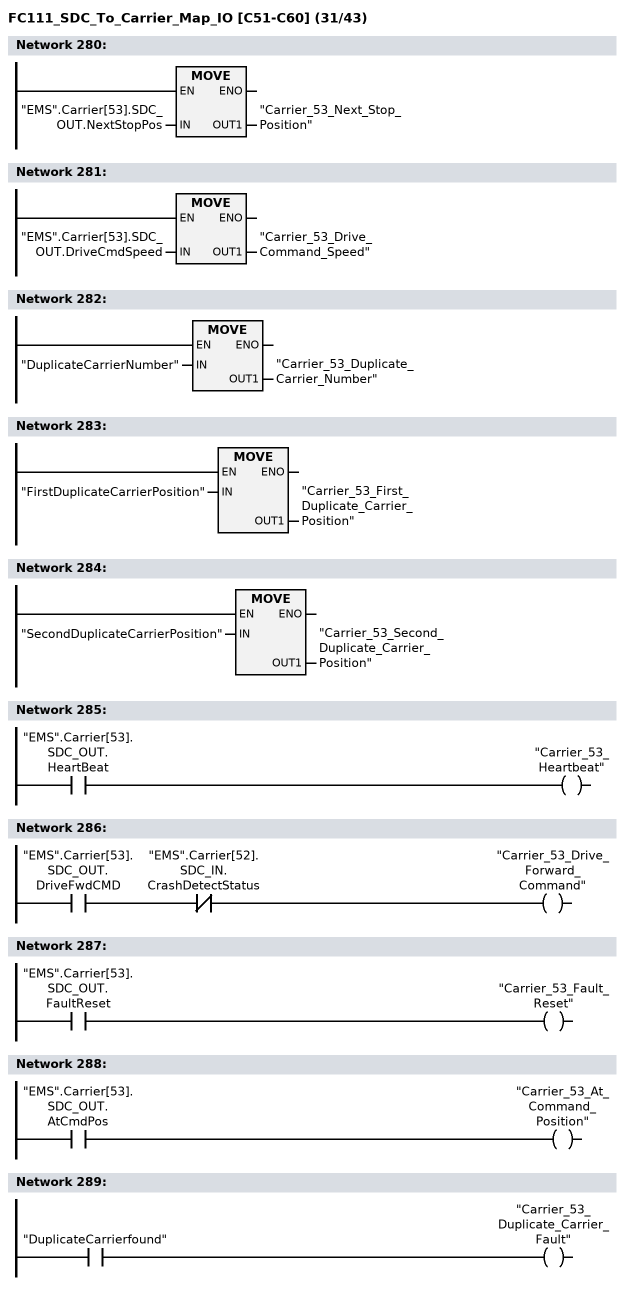
   RUNG wire#powerrail
      Move(in := "EMS".Carrier[53].SDC_OUT.NextStopPos, out1 => "Carrier_53_Next_Stop_Position")
   END_RUNG
   // the same network as SCL:
   "Carrier_53_Next_Stop_Position" := "EMS".Carrier[53].SDC_OUT.NextStopPos;
END_REGION

REGION Network 281
   RUNG wire#powerrail
      Move(in := "EMS".Carrier[53].SDC_OUT.DriveCmdSpeed, out1 => "Carrier_53_Drive_Command_Speed")
   END_RUNG
   // the same network as SCL:
   "Carrier_53_Drive_Command_Speed" := "EMS".Carrier[53].SDC_OUT.DriveCmdSpeed;
END_REGION

REGION Network 282
   RUNG wire#powerrail
      Move(in := "DuplicateCarrierNumber", out1 => "Carrier_53_Duplicate_Carrier_Number")
   END_RUNG
   // the same network as SCL:
   "Carrier_53_Duplicate_Carrier_Number" := "DuplicateCarrierNumber";
END_REGION

REGION Network 283
   RUNG wire#powerrail
      Move(in := "FirstDuplicateCarrierPosition", out1 => "Carrier_53_First_Duplicate_Carrier_Position")
   END_RUNG
   // the same network as SCL:
   "Carrier_53_First_Duplicate_Carrier_Position" := "FirstDuplicateCarrierPosition";
END_REGION

REGION Network 284
   RUNG wire#powerrail
      Move(in := "SecondDuplicateCarrierPosition", out1 => "Carrier_53_Second_Duplicate_Carrier_Position")
   END_RUNG
   // the same network as SCL:
   "Carrier_53_Second_Duplicate_Carrier_Position" := "SecondDuplicateCarrierPosition";
END_REGION

REGION Network 285
   RUNG wire#powerrail
      Contact( "EMS".Carrier[53].SDC_OUT.HeartBeat )
      Coil( "Carrier_53_Heartbeat" )
   END_RUNG
   // the same network as SCL:
   "Carrier_53_Heartbeat" := "EMS".Carrier[53].SDC_OUT.HeartBeat;
END_REGION

REGION Network 286
   RUNG wire#powerrail
      Contact( "EMS".Carrier[53].SDC_OUT.DriveFwdCMD )
      I_Contact( "EMS".Carrier[52].SDC_IN.CrashDetectStatus )
      Coil( "Carrier_53_Drive_Forward_Command" )
   END_RUNG
   // the same network as SCL:
   "Carrier_53_Drive_Forward_Command" := "EMS".Carrier[53].SDC_OUT.DriveFwdCMD AND NOT "EMS".Carrier[52].SDC_IN.CrashDetectStatus;
END_REGION

REGION Network 287
   RUNG wire#powerrail
      Contact( "EMS".Carrier[53].SDC_OUT.FaultReset )
      Coil( "Carrier_53_Fault_Reset" )
   END_RUNG
   // the same network as SCL:
   "Carrier_53_Fault_Reset" := "EMS".Carrier[53].SDC_OUT.FaultReset;
END_REGION

REGION Network 288
   RUNG wire#powerrail
      Contact( "EMS".Carrier[53].SDC_OUT.AtCmdPos )
      Coil( "Carrier_53_At_Command_Position" )
   END_RUNG
   // the same network as SCL:
   "Carrier_53_At_Command_Position" := "EMS".Carrier[53].SDC_OUT.AtCmdPos;
END_REGION

REGION Network 289
   RUNG wire#powerrail
      Contact( "DuplicateCarrierfound" )
      Coil( "Carrier_53_Duplicate_Carrier_Fault" )
   END_RUNG
   // the same network as SCL:
   "Carrier_53_Duplicate_Carrier_Fault" := "DuplicateCarrierfound";
END_REGION

REGION Network 290
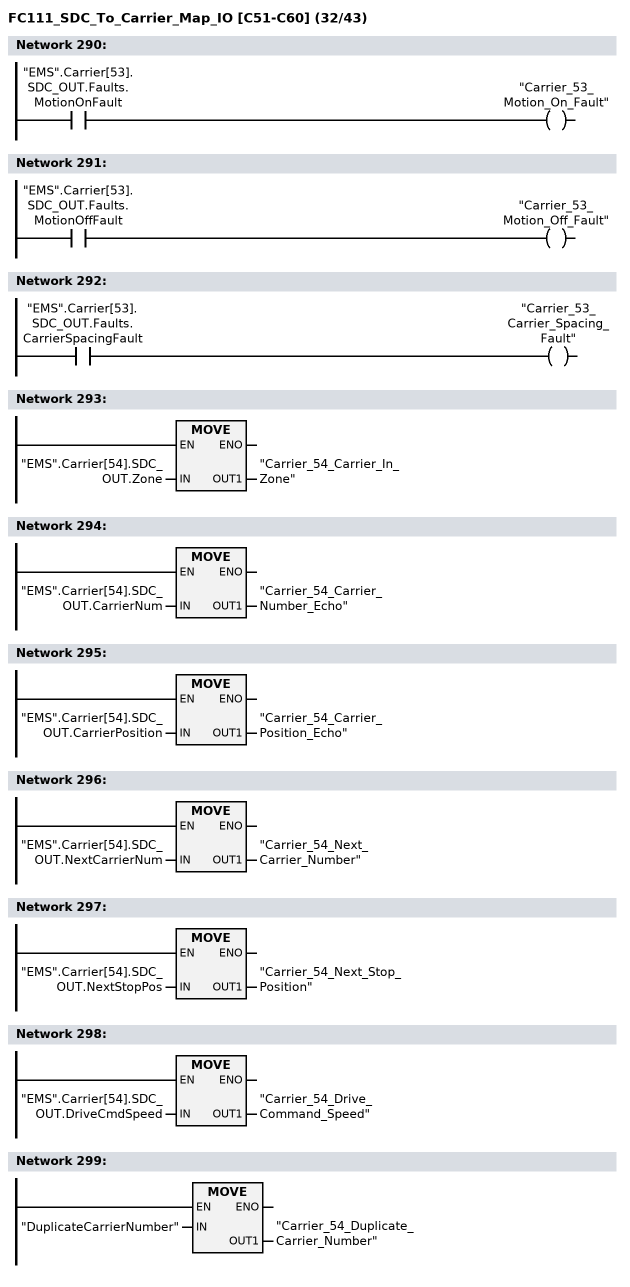
   RUNG wire#powerrail
      Contact( "EMS".Carrier[53].SDC_OUT.Faults.MotionOnFault )
      Coil( "Carrier_53_Motion_On_Fault" )
   END_RUNG
   // the same network as SCL:
   "Carrier_53_Motion_On_Fault" := "EMS".Carrier[53].SDC_OUT.Faults.MotionOnFault;
END_REGION

REGION Network 291
   RUNG wire#powerrail
      Contact( "EMS".Carrier[53].SDC_OUT.Faults.MotionOffFault )
      Coil( "Carrier_53_Motion_Off_Fault" )
   END_RUNG
   // the same network as SCL:
   "Carrier_53_Motion_Off_Fault" := "EMS".Carrier[53].SDC_OUT.Faults.MotionOffFault;
END_REGION

REGION Network 292
   RUNG wire#powerrail
      Contact( "EMS".Carrier[53].SDC_OUT.Faults.CarrierSpacingFault )
      Coil( "Carrier_53_Carrier_Spacing_Fault" )
   END_RUNG
   // the same network as SCL:
   "Carrier_53_Carrier_Spacing_Fault" := "EMS".Carrier[53].SDC_OUT.Faults.CarrierSpacingFault;
END_REGION

REGION Network 293
   RUNG wire#powerrail
      Move(in := "EMS".Carrier[54].SDC_OUT.Zone, out1 => "Carrier_54_Carrier_In_Zone")
   END_RUNG
   // the same network as SCL:
   "Carrier_54_Carrier_In_Zone" := "EMS".Carrier[54].SDC_OUT.Zone;
END_REGION

REGION Network 294
   RUNG wire#powerrail
      Move(in := "EMS".Carrier[54].SDC_OUT.CarrierNum, out1 => "Carrier_54_Carrier_Number_Echo")
   END_RUNG
   // the same network as SCL:
   "Carrier_54_Carrier_Number_Echo" := "EMS".Carrier[54].SDC_OUT.CarrierNum;
END_REGION

REGION Network 295
   RUNG wire#powerrail
      Move(in := "EMS".Carrier[54].SDC_OUT.CarrierPosition, out1 => "Carrier_54_Carrier_Position_Echo")
   END_RUNG
   // the same network as SCL:
   "Carrier_54_Carrier_Position_Echo" := "EMS".Carrier[54].SDC_OUT.CarrierPosition;
END_REGION

REGION Network 296
   RUNG wire#powerrail
      Move(in := "EMS".Carrier[54].SDC_OUT.NextCarrierNum, out1 => "Carrier_54_Next_Carrier_Number")
   END_RUNG
   // the same network as SCL:
   "Carrier_54_Next_Carrier_Number" := "EMS".Carrier[54].SDC_OUT.NextCarrierNum;
END_REGION

REGION Network 297
   RUNG wire#powerrail
      Move(in := "EMS".Carrier[54].SDC_OUT.NextStopPos, out1 => "Carrier_54_Next_Stop_Position")
   END_RUNG
   // the same network as SCL:
   "Carrier_54_Next_Stop_Position" := "EMS".Carrier[54].SDC_OUT.NextStopPos;
END_REGION

REGION Network 298
   RUNG wire#powerrail
      Move(in := "EMS".Carrier[54].SDC_OUT.DriveCmdSpeed, out1 => "Carrier_54_Drive_Command_Speed")
   END_RUNG
   // the same network as SCL:
   "Carrier_54_Drive_Command_Speed" := "EMS".Carrier[54].SDC_OUT.DriveCmdSpeed;
END_REGION

REGION Network 299
   RUNG wire#powerrail
      Move(in := "DuplicateCarrierNumber", out1 => "Carrier_54_Duplicate_Carrier_Number")
   END_RUNG
   // the same network as SCL:
   "Carrier_54_Duplicate_Carrier_Number" := "DuplicateCarrierNumber";
END_REGION

REGION Network 300
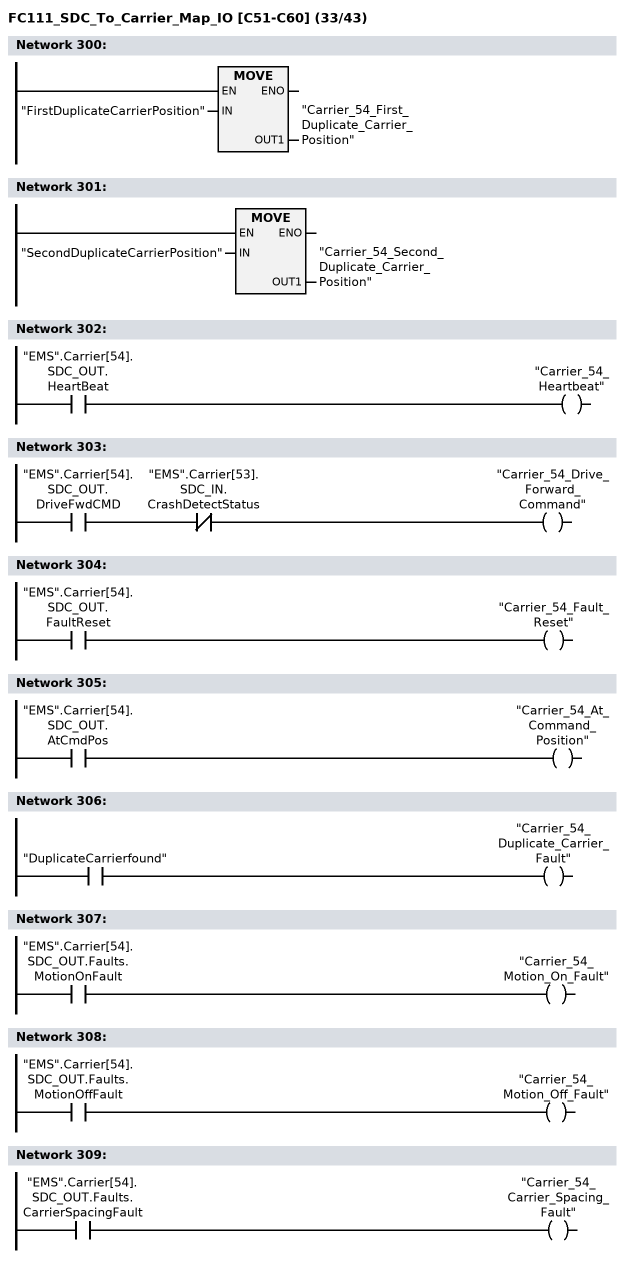
   RUNG wire#powerrail
      Move(in := "FirstDuplicateCarrierPosition", out1 => "Carrier_54_First_Duplicate_Carrier_Position")
   END_RUNG
   // the same network as SCL:
   "Carrier_54_First_Duplicate_Carrier_Position" := "FirstDuplicateCarrierPosition";
END_REGION

REGION Network 301
   RUNG wire#powerrail
      Move(in := "SecondDuplicateCarrierPosition", out1 => "Carrier_54_Second_Duplicate_Carrier_Position")
   END_RUNG
   // the same network as SCL:
   "Carrier_54_Second_Duplicate_Carrier_Position" := "SecondDuplicateCarrierPosition";
END_REGION

REGION Network 302
   RUNG wire#powerrail
      Contact( "EMS".Carrier[54].SDC_OUT.HeartBeat )
      Coil( "Carrier_54_Heartbeat" )
   END_RUNG
   // the same network as SCL:
   "Carrier_54_Heartbeat" := "EMS".Carrier[54].SDC_OUT.HeartBeat;
END_REGION

REGION Network 303
   RUNG wire#powerrail
      Contact( "EMS".Carrier[54].SDC_OUT.DriveFwdCMD )
      I_Contact( "EMS".Carrier[53].SDC_IN.CrashDetectStatus )
      Coil( "Carrier_54_Drive_Forward_Command" )
   END_RUNG
   // the same network as SCL:
   "Carrier_54_Drive_Forward_Command" := "EMS".Carrier[54].SDC_OUT.DriveFwdCMD AND NOT "EMS".Carrier[53].SDC_IN.CrashDetectStatus;
END_REGION

REGION Network 304
   RUNG wire#powerrail
      Contact( "EMS".Carrier[54].SDC_OUT.FaultReset )
      Coil( "Carrier_54_Fault_Reset" )
   END_RUNG
   // the same network as SCL:
   "Carrier_54_Fault_Reset" := "EMS".Carrier[54].SDC_OUT.FaultReset;
END_REGION

REGION Network 305
   RUNG wire#powerrail
      Contact( "EMS".Carrier[54].SDC_OUT.AtCmdPos )
      Coil( "Carrier_54_At_Command_Position" )
   END_RUNG
   // the same network as SCL:
   "Carrier_54_At_Command_Position" := "EMS".Carrier[54].SDC_OUT.AtCmdPos;
END_REGION

REGION Network 306
   RUNG wire#powerrail
      Contact( "DuplicateCarrierfound" )
      Coil( "Carrier_54_Duplicate_Carrier_Fault" )
   END_RUNG
   // the same network as SCL:
   "Carrier_54_Duplicate_Carrier_Fault" := "DuplicateCarrierfound";
END_REGION

REGION Network 307
   RUNG wire#powerrail
      Contact( "EMS".Carrier[54].SDC_OUT.Faults.MotionOnFault )
      Coil( "Carrier_54_Motion_On_Fault" )
   END_RUNG
   // the same network as SCL:
   "Carrier_54_Motion_On_Fault" := "EMS".Carrier[54].SDC_OUT.Faults.MotionOnFault;
END_REGION

REGION Network 308
   RUNG wire#powerrail
      Contact( "EMS".Carrier[54].SDC_OUT.Faults.MotionOffFault )
      Coil( "Carrier_54_Motion_Off_Fault" )
   END_RUNG
   // the same network as SCL:
   "Carrier_54_Motion_Off_Fault" := "EMS".Carrier[54].SDC_OUT.Faults.MotionOffFault;
END_REGION

REGION Network 309
   RUNG wire#powerrail
      Contact( "EMS".Carrier[54].SDC_OUT.Faults.CarrierSpacingFault )
      Coil( "Carrier_54_Carrier_Spacing_Fault" )
   END_RUNG
   // the same network as SCL:
   "Carrier_54_Carrier_Spacing_Fault" := "EMS".Carrier[54].SDC_OUT.Faults.CarrierSpacingFault;
END_REGION

REGION Network 310
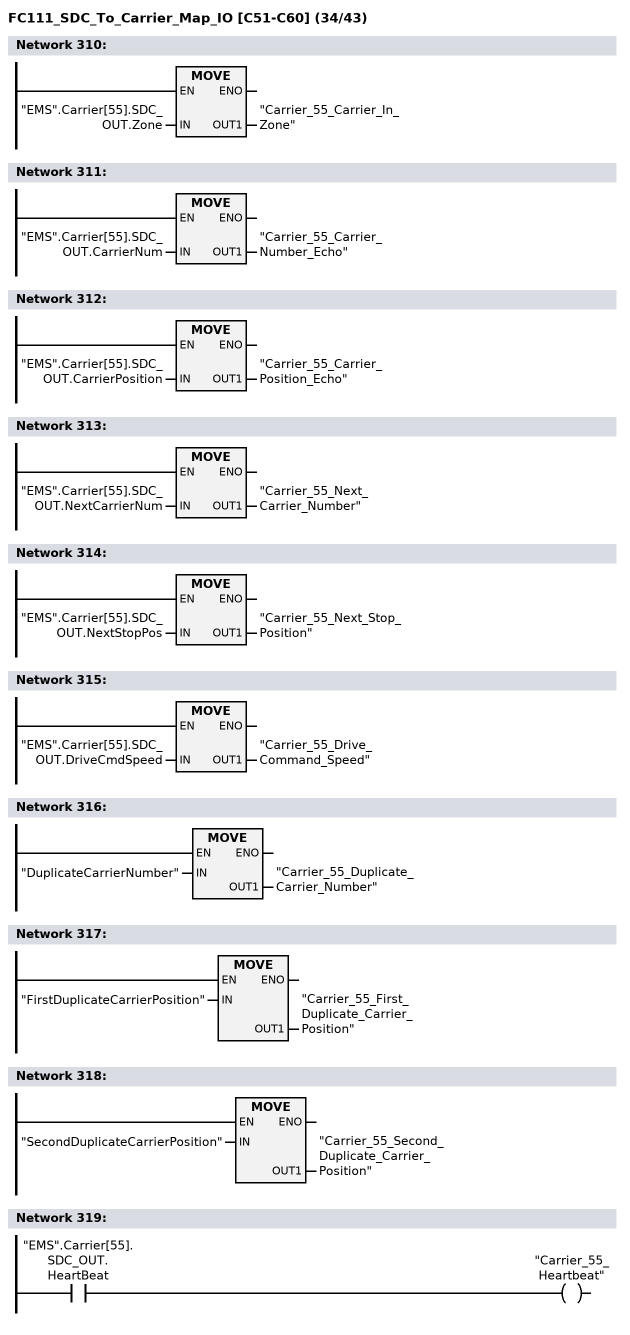
   RUNG wire#powerrail
      Move(in := "EMS".Carrier[55].SDC_OUT.Zone, out1 => "Carrier_55_Carrier_In_Zone")
   END_RUNG
   // the same network as SCL:
   "Carrier_55_Carrier_In_Zone" := "EMS".Carrier[55].SDC_OUT.Zone;
END_REGION

REGION Network 311
   RUNG wire#powerrail
      Move(in := "EMS".Carrier[55].SDC_OUT.CarrierNum, out1 => "Carrier_55_Carrier_Number_Echo")
   END_RUNG
   // the same network as SCL:
   "Carrier_55_Carrier_Number_Echo" := "EMS".Carrier[55].SDC_OUT.CarrierNum;
END_REGION

REGION Network 312
   RUNG wire#powerrail
      Move(in := "EMS".Carrier[55].SDC_OUT.CarrierPosition, out1 => "Carrier_55_Carrier_Position_Echo")
   END_RUNG
   // the same network as SCL:
   "Carrier_55_Carrier_Position_Echo" := "EMS".Carrier[55].SDC_OUT.CarrierPosition;
END_REGION

REGION Network 313
   RUNG wire#powerrail
      Move(in := "EMS".Carrier[55].SDC_OUT.NextCarrierNum, out1 => "Carrier_55_Next_Carrier_Number")
   END_RUNG
   // the same network as SCL:
   "Carrier_55_Next_Carrier_Number" := "EMS".Carrier[55].SDC_OUT.NextCarrierNum;
END_REGION

REGION Network 314
   RUNG wire#powerrail
      Move(in := "EMS".Carrier[55].SDC_OUT.NextStopPos, out1 => "Carrier_55_Next_Stop_Position")
   END_RUNG
   // the same network as SCL:
   "Carrier_55_Next_Stop_Position" := "EMS".Carrier[55].SDC_OUT.NextStopPos;
END_REGION

REGION Network 315
   RUNG wire#powerrail
      Move(in := "EMS".Carrier[55].SDC_OUT.DriveCmdSpeed, out1 => "Carrier_55_Drive_Command_Speed")
   END_RUNG
   // the same network as SCL:
   "Carrier_55_Drive_Command_Speed" := "EMS".Carrier[55].SDC_OUT.DriveCmdSpeed;
END_REGION

REGION Network 316
   RUNG wire#powerrail
      Move(in := "DuplicateCarrierNumber", out1 => "Carrier_55_Duplicate_Carrier_Number")
   END_RUNG
   // the same network as SCL:
   "Carrier_55_Duplicate_Carrier_Number" := "DuplicateCarrierNumber";
END_REGION

REGION Network 317
   RUNG wire#powerrail
      Move(in := "FirstDuplicateCarrierPosition", out1 => "Carrier_55_First_Duplicate_Carrier_Position")
   END_RUNG
   // the same network as SCL:
   "Carrier_55_First_Duplicate_Carrier_Position" := "FirstDuplicateCarrierPosition";
END_REGION

REGION Network 318
   RUNG wire#powerrail
      Move(in := "SecondDuplicateCarrierPosition", out1 => "Carrier_55_Second_Duplicate_Carrier_Position")
   END_RUNG
   // the same network as SCL:
   "Carrier_55_Second_Duplicate_Carrier_Position" := "SecondDuplicateCarrierPosition";
END_REGION

REGION Network 319
   RUNG wire#powerrail
      Contact( "EMS".Carrier[55].SDC_OUT.HeartBeat )
      Coil( "Carrier_55_Heartbeat" )
   END_RUNG
   // the same network as SCL:
   "Carrier_55_Heartbeat" := "EMS".Carrier[55].SDC_OUT.HeartBeat;
END_REGION

REGION Network 320
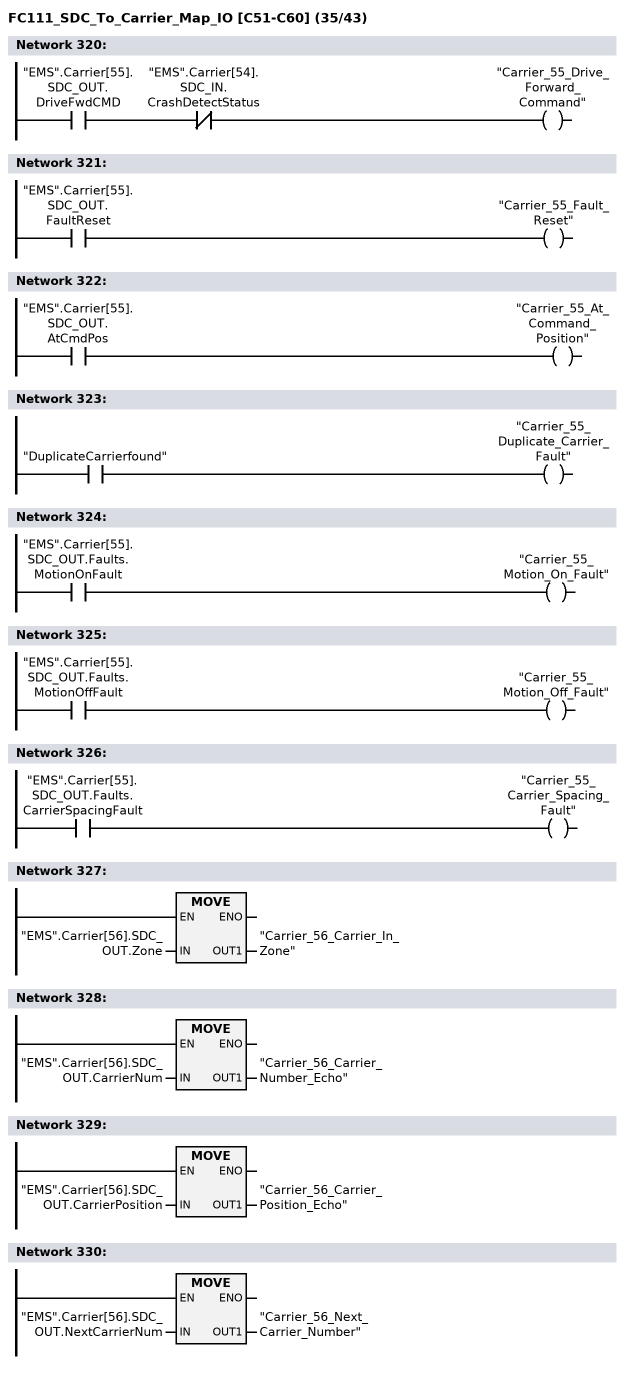
   RUNG wire#powerrail
      Contact( "EMS".Carrier[55].SDC_OUT.DriveFwdCMD )
      I_Contact( "EMS".Carrier[54].SDC_IN.CrashDetectStatus )
      Coil( "Carrier_55_Drive_Forward_Command" )
   END_RUNG
   // the same network as SCL:
   "Carrier_55_Drive_Forward_Command" := "EMS".Carrier[55].SDC_OUT.DriveFwdCMD AND NOT "EMS".Carrier[54].SDC_IN.CrashDetectStatus;
END_REGION

REGION Network 321
   RUNG wire#powerrail
      Contact( "EMS".Carrier[55].SDC_OUT.FaultReset )
      Coil( "Carrier_55_Fault_Reset" )
   END_RUNG
   // the same network as SCL:
   "Carrier_55_Fault_Reset" := "EMS".Carrier[55].SDC_OUT.FaultReset;
END_REGION

REGION Network 322
   RUNG wire#powerrail
      Contact( "EMS".Carrier[55].SDC_OUT.AtCmdPos )
      Coil( "Carrier_55_At_Command_Position" )
   END_RUNG
   // the same network as SCL:
   "Carrier_55_At_Command_Position" := "EMS".Carrier[55].SDC_OUT.AtCmdPos;
END_REGION

REGION Network 323
   RUNG wire#powerrail
      Contact( "DuplicateCarrierfound" )
      Coil( "Carrier_55_Duplicate_Carrier_Fault" )
   END_RUNG
   // the same network as SCL:
   "Carrier_55_Duplicate_Carrier_Fault" := "DuplicateCarrierfound";
END_REGION

REGION Network 324
   RUNG wire#powerrail
      Contact( "EMS".Carrier[55].SDC_OUT.Faults.MotionOnFault )
      Coil( "Carrier_55_Motion_On_Fault" )
   END_RUNG
   // the same network as SCL:
   "Carrier_55_Motion_On_Fault" := "EMS".Carrier[55].SDC_OUT.Faults.MotionOnFault;
END_REGION

REGION Network 325
   RUNG wire#powerrail
      Contact( "EMS".Carrier[55].SDC_OUT.Faults.MotionOffFault )
      Coil( "Carrier_55_Motion_Off_Fault" )
   END_RUNG
   // the same network as SCL:
   "Carrier_55_Motion_Off_Fault" := "EMS".Carrier[55].SDC_OUT.Faults.MotionOffFault;
END_REGION

REGION Network 326
   RUNG wire#powerrail
      Contact( "EMS".Carrier[55].SDC_OUT.Faults.CarrierSpacingFault )
      Coil( "Carrier_55_Carrier_Spacing_Fault" )
   END_RUNG
   // the same network as SCL:
   "Carrier_55_Carrier_Spacing_Fault" := "EMS".Carrier[55].SDC_OUT.Faults.CarrierSpacingFault;
END_REGION

REGION Network 327
   RUNG wire#powerrail
      Move(in := "EMS".Carrier[56].SDC_OUT.Zone, out1 => "Carrier_56_Carrier_In_Zone")
   END_RUNG
   // the same network as SCL:
   "Carrier_56_Carrier_In_Zone" := "EMS".Carrier[56].SDC_OUT.Zone;
END_REGION

REGION Network 328
   RUNG wire#powerrail
      Move(in := "EMS".Carrier[56].SDC_OUT.CarrierNum, out1 => "Carrier_56_Carrier_Number_Echo")
   END_RUNG
   // the same network as SCL:
   "Carrier_56_Carrier_Number_Echo" := "EMS".Carrier[56].SDC_OUT.CarrierNum;
END_REGION

REGION Network 329
   RUNG wire#powerrail
      Move(in := "EMS".Carrier[56].SDC_OUT.CarrierPosition, out1 => "Carrier_56_Carrier_Position_Echo")
   END_RUNG
   // the same network as SCL:
   "Carrier_56_Carrier_Position_Echo" := "EMS".Carrier[56].SDC_OUT.CarrierPosition;
END_REGION

REGION Network 330
   RUNG wire#powerrail
      Move(in := "EMS".Carrier[56].SDC_OUT.NextCarrierNum, out1 => "Carrier_56_Next_Carrier_Number")
   END_RUNG
   // the same network as SCL:
   "Carrier_56_Next_Carrier_Number" := "EMS".Carrier[56].SDC_OUT.NextCarrierNum;
END_REGION

REGION Network 331
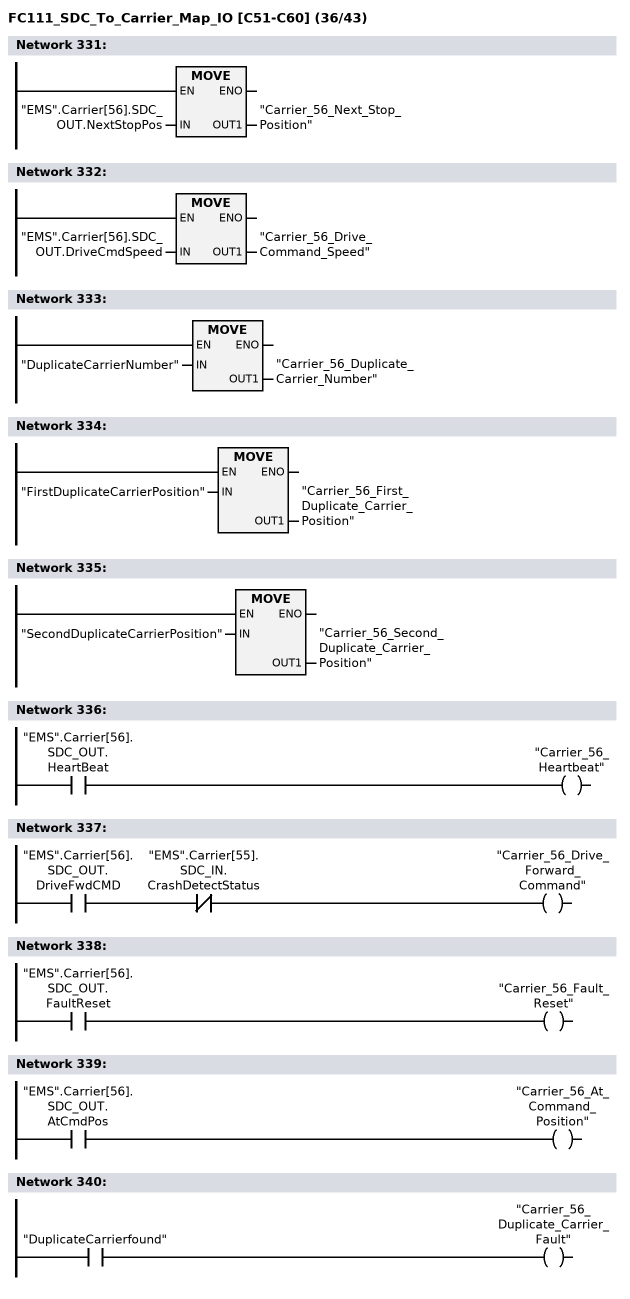
   RUNG wire#powerrail
      Move(in := "EMS".Carrier[56].SDC_OUT.NextStopPos, out1 => "Carrier_56_Next_Stop_Position")
   END_RUNG
   // the same network as SCL:
   "Carrier_56_Next_Stop_Position" := "EMS".Carrier[56].SDC_OUT.NextStopPos;
END_REGION

REGION Network 332
   RUNG wire#powerrail
      Move(in := "EMS".Carrier[56].SDC_OUT.DriveCmdSpeed, out1 => "Carrier_56_Drive_Command_Speed")
   END_RUNG
   // the same network as SCL:
   "Carrier_56_Drive_Command_Speed" := "EMS".Carrier[56].SDC_OUT.DriveCmdSpeed;
END_REGION

REGION Network 333
   RUNG wire#powerrail
      Move(in := "DuplicateCarrierNumber", out1 => "Carrier_56_Duplicate_Carrier_Number")
   END_RUNG
   // the same network as SCL:
   "Carrier_56_Duplicate_Carrier_Number" := "DuplicateCarrierNumber";
END_REGION

REGION Network 334
   RUNG wire#powerrail
      Move(in := "FirstDuplicateCarrierPosition", out1 => "Carrier_56_First_Duplicate_Carrier_Position")
   END_RUNG
   // the same network as SCL:
   "Carrier_56_First_Duplicate_Carrier_Position" := "FirstDuplicateCarrierPosition";
END_REGION

REGION Network 335
   RUNG wire#powerrail
      Move(in := "SecondDuplicateCarrierPosition", out1 => "Carrier_56_Second_Duplicate_Carrier_Position")
   END_RUNG
   // the same network as SCL:
   "Carrier_56_Second_Duplicate_Carrier_Position" := "SecondDuplicateCarrierPosition";
END_REGION

REGION Network 336
   RUNG wire#powerrail
      Contact( "EMS".Carrier[56].SDC_OUT.HeartBeat )
      Coil( "Carrier_56_Heartbeat" )
   END_RUNG
   // the same network as SCL:
   "Carrier_56_Heartbeat" := "EMS".Carrier[56].SDC_OUT.HeartBeat;
END_REGION

REGION Network 337
   RUNG wire#powerrail
      Contact( "EMS".Carrier[56].SDC_OUT.DriveFwdCMD )
      I_Contact( "EMS".Carrier[55].SDC_IN.CrashDetectStatus )
      Coil( "Carrier_56_Drive_Forward_Command" )
   END_RUNG
   // the same network as SCL:
   "Carrier_56_Drive_Forward_Command" := "EMS".Carrier[56].SDC_OUT.DriveFwdCMD AND NOT "EMS".Carrier[55].SDC_IN.CrashDetectStatus;
END_REGION

REGION Network 338
   RUNG wire#powerrail
      Contact( "EMS".Carrier[56].SDC_OUT.FaultReset )
      Coil( "Carrier_56_Fault_Reset" )
   END_RUNG
   // the same network as SCL:
   "Carrier_56_Fault_Reset" := "EMS".Carrier[56].SDC_OUT.FaultReset;
END_REGION

REGION Network 339
   RUNG wire#powerrail
      Contact( "EMS".Carrier[56].SDC_OUT.AtCmdPos )
      Coil( "Carrier_56_At_Command_Position" )
   END_RUNG
   // the same network as SCL:
   "Carrier_56_At_Command_Position" := "EMS".Carrier[56].SDC_OUT.AtCmdPos;
END_REGION

REGION Network 340
   RUNG wire#powerrail
      Contact( "DuplicateCarrierfound" )
      Coil( "Carrier_56_Duplicate_Carrier_Fault" )
   END_RUNG
   // the same network as SCL:
   "Carrier_56_Duplicate_Carrier_Fault" := "DuplicateCarrierfound";
END_REGION

REGION Network 341
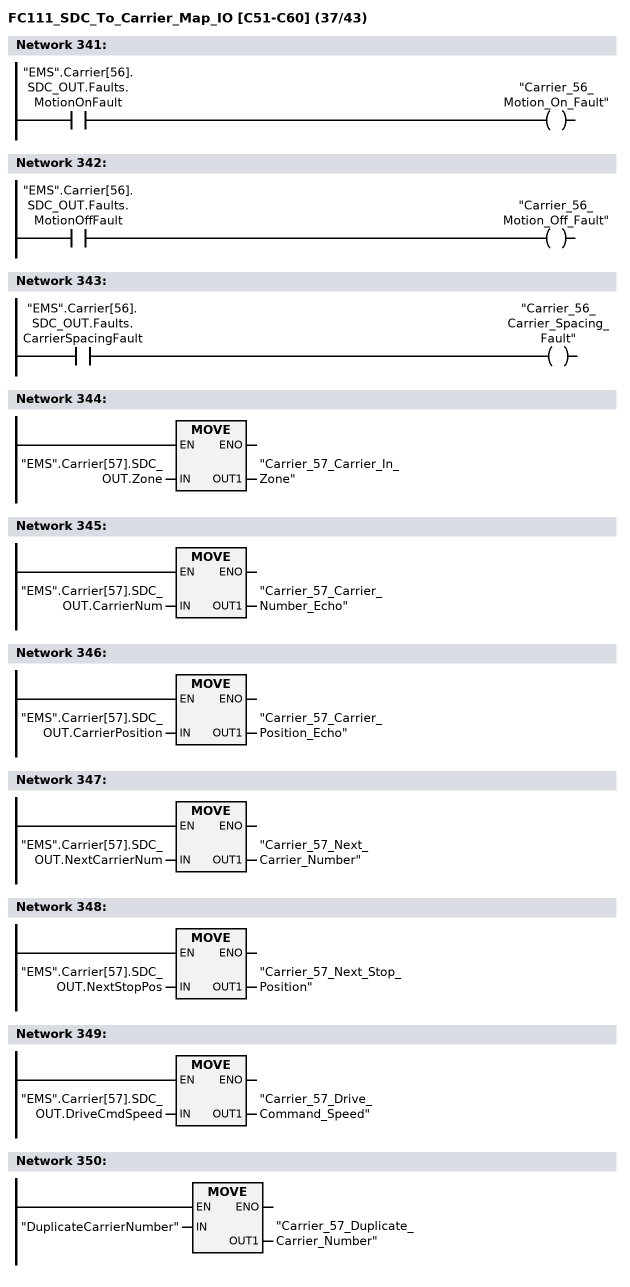
   RUNG wire#powerrail
      Contact( "EMS".Carrier[56].SDC_OUT.Faults.MotionOnFault )
      Coil( "Carrier_56_Motion_On_Fault" )
   END_RUNG
   // the same network as SCL:
   "Carrier_56_Motion_On_Fault" := "EMS".Carrier[56].SDC_OUT.Faults.MotionOnFault;
END_REGION

REGION Network 342
   RUNG wire#powerrail
      Contact( "EMS".Carrier[56].SDC_OUT.Faults.MotionOffFault )
      Coil( "Carrier_56_Motion_Off_Fault" )
   END_RUNG
   // the same network as SCL:
   "Carrier_56_Motion_Off_Fault" := "EMS".Carrier[56].SDC_OUT.Faults.MotionOffFault;
END_REGION

REGION Network 343
   RUNG wire#powerrail
      Contact( "EMS".Carrier[56].SDC_OUT.Faults.CarrierSpacingFault )
      Coil( "Carrier_56_Carrier_Spacing_Fault" )
   END_RUNG
   // the same network as SCL:
   "Carrier_56_Carrier_Spacing_Fault" := "EMS".Carrier[56].SDC_OUT.Faults.CarrierSpacingFault;
END_REGION

REGION Network 344
   RUNG wire#powerrail
      Move(in := "EMS".Carrier[57].SDC_OUT.Zone, out1 => "Carrier_57_Carrier_In_Zone")
   END_RUNG
   // the same network as SCL:
   "Carrier_57_Carrier_In_Zone" := "EMS".Carrier[57].SDC_OUT.Zone;
END_REGION

REGION Network 345
   RUNG wire#powerrail
      Move(in := "EMS".Carrier[57].SDC_OUT.CarrierNum, out1 => "Carrier_57_Carrier_Number_Echo")
   END_RUNG
   // the same network as SCL:
   "Carrier_57_Carrier_Number_Echo" := "EMS".Carrier[57].SDC_OUT.CarrierNum;
END_REGION

REGION Network 346
   RUNG wire#powerrail
      Move(in := "EMS".Carrier[57].SDC_OUT.CarrierPosition, out1 => "Carrier_57_Carrier_Position_Echo")
   END_RUNG
   // the same network as SCL:
   "Carrier_57_Carrier_Position_Echo" := "EMS".Carrier[57].SDC_OUT.CarrierPosition;
END_REGION

REGION Network 347
   RUNG wire#powerrail
      Move(in := "EMS".Carrier[57].SDC_OUT.NextCarrierNum, out1 => "Carrier_57_Next_Carrier_Number")
   END_RUNG
   // the same network as SCL:
   "Carrier_57_Next_Carrier_Number" := "EMS".Carrier[57].SDC_OUT.NextCarrierNum;
END_REGION

REGION Network 348
   RUNG wire#powerrail
      Move(in := "EMS".Carrier[57].SDC_OUT.NextStopPos, out1 => "Carrier_57_Next_Stop_Position")
   END_RUNG
   // the same network as SCL:
   "Carrier_57_Next_Stop_Position" := "EMS".Carrier[57].SDC_OUT.NextStopPos;
END_REGION

REGION Network 349
   RUNG wire#powerrail
      Move(in := "EMS".Carrier[57].SDC_OUT.DriveCmdSpeed, out1 => "Carrier_57_Drive_Command_Speed")
   END_RUNG
   // the same network as SCL:
   "Carrier_57_Drive_Command_Speed" := "EMS".Carrier[57].SDC_OUT.DriveCmdSpeed;
END_REGION

REGION Network 350
   RUNG wire#powerrail
      Move(in := "DuplicateCarrierNumber", out1 => "Carrier_57_Duplicate_Carrier_Number")
   END_RUNG
   // the same network as SCL:
   "Carrier_57_Duplicate_Carrier_Number" := "DuplicateCarrierNumber";
END_REGION

REGION Network 351
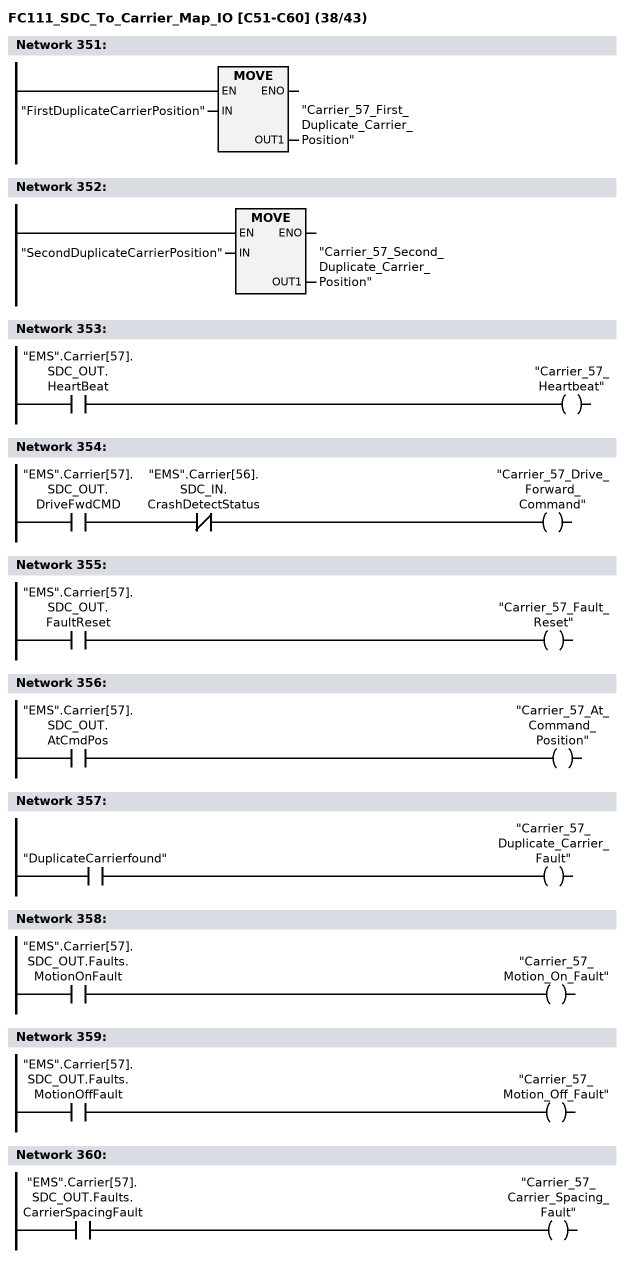
   RUNG wire#powerrail
      Move(in := "FirstDuplicateCarrierPosition", out1 => "Carrier_57_First_Duplicate_Carrier_Position")
   END_RUNG
   // the same network as SCL:
   "Carrier_57_First_Duplicate_Carrier_Position" := "FirstDuplicateCarrierPosition";
END_REGION

REGION Network 352
   RUNG wire#powerrail
      Move(in := "SecondDuplicateCarrierPosition", out1 => "Carrier_57_Second_Duplicate_Carrier_Position")
   END_RUNG
   // the same network as SCL:
   "Carrier_57_Second_Duplicate_Carrier_Position" := "SecondDuplicateCarrierPosition";
END_REGION

REGION Network 353
   RUNG wire#powerrail
      Contact( "EMS".Carrier[57].SDC_OUT.HeartBeat )
      Coil( "Carrier_57_Heartbeat" )
   END_RUNG
   // the same network as SCL:
   "Carrier_57_Heartbeat" := "EMS".Carrier[57].SDC_OUT.HeartBeat;
END_REGION

REGION Network 354
   RUNG wire#powerrail
      Contact( "EMS".Carrier[57].SDC_OUT.DriveFwdCMD )
      I_Contact( "EMS".Carrier[56].SDC_IN.CrashDetectStatus )
      Coil( "Carrier_57_Drive_Forward_Command" )
   END_RUNG
   // the same network as SCL:
   "Carrier_57_Drive_Forward_Command" := "EMS".Carrier[57].SDC_OUT.DriveFwdCMD AND NOT "EMS".Carrier[56].SDC_IN.CrashDetectStatus;
END_REGION

REGION Network 355
   RUNG wire#powerrail
      Contact( "EMS".Carrier[57].SDC_OUT.FaultReset )
      Coil( "Carrier_57_Fault_Reset" )
   END_RUNG
   // the same network as SCL:
   "Carrier_57_Fault_Reset" := "EMS".Carrier[57].SDC_OUT.FaultReset;
END_REGION

REGION Network 356
   RUNG wire#powerrail
      Contact( "EMS".Carrier[57].SDC_OUT.AtCmdPos )
      Coil( "Carrier_57_At_Command_Position" )
   END_RUNG
   // the same network as SCL:
   "Carrier_57_At_Command_Position" := "EMS".Carrier[57].SDC_OUT.AtCmdPos;
END_REGION

REGION Network 357
   RUNG wire#powerrail
      Contact( "DuplicateCarrierfound" )
      Coil( "Carrier_57_Duplicate_Carrier_Fault" )
   END_RUNG
   // the same network as SCL:
   "Carrier_57_Duplicate_Carrier_Fault" := "DuplicateCarrierfound";
END_REGION

REGION Network 358
   RUNG wire#powerrail
      Contact( "EMS".Carrier[57].SDC_OUT.Faults.MotionOnFault )
      Coil( "Carrier_57_Motion_On_Fault" )
   END_RUNG
   // the same network as SCL:
   "Carrier_57_Motion_On_Fault" := "EMS".Carrier[57].SDC_OUT.Faults.MotionOnFault;
END_REGION

REGION Network 359
   RUNG wire#powerrail
      Contact( "EMS".Carrier[57].SDC_OUT.Faults.MotionOffFault )
      Coil( "Carrier_57_Motion_Off_Fault" )
   END_RUNG
   // the same network as SCL:
   "Carrier_57_Motion_Off_Fault" := "EMS".Carrier[57].SDC_OUT.Faults.MotionOffFault;
END_REGION

REGION Network 360
   RUNG wire#powerrail
      Contact( "EMS".Carrier[57].SDC_OUT.Faults.CarrierSpacingFault )
      Coil( "Carrier_57_Carrier_Spacing_Fault" )
   END_RUNG
   // the same network as SCL:
   "Carrier_57_Carrier_Spacing_Fault" := "EMS".Carrier[57].SDC_OUT.Faults.CarrierSpacingFault;
END_REGION

REGION Network 361
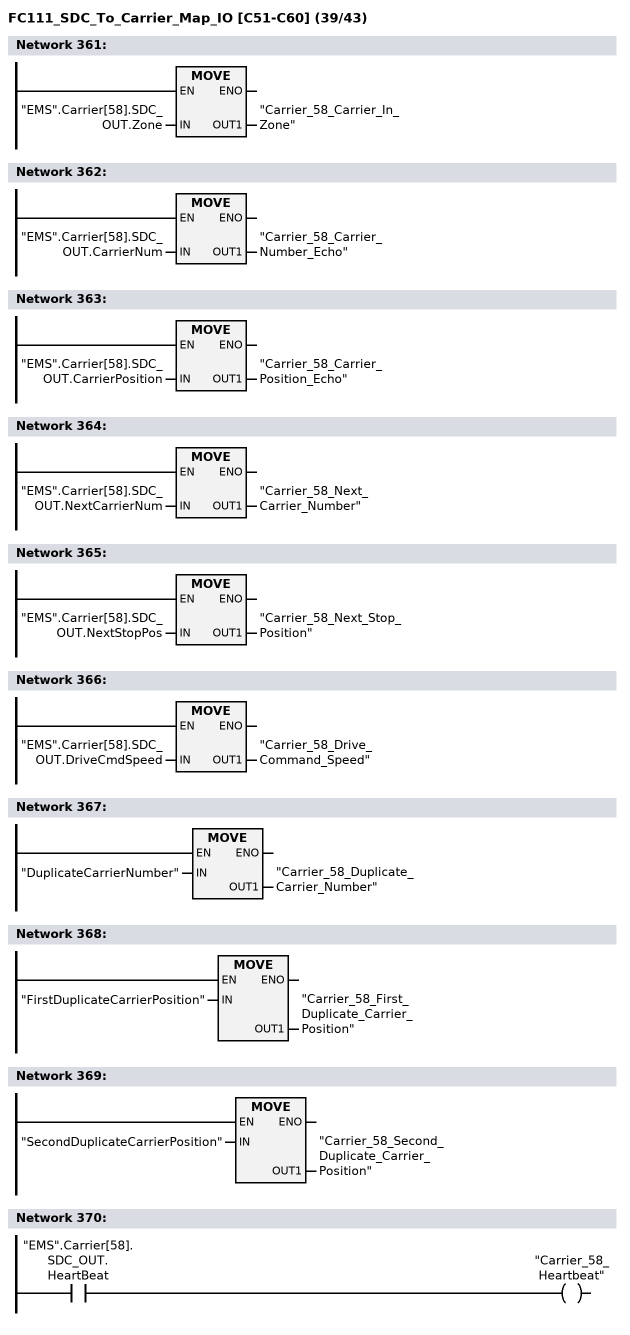
   RUNG wire#powerrail
      Move(in := "EMS".Carrier[58].SDC_OUT.Zone, out1 => "Carrier_58_Carrier_In_Zone")
   END_RUNG
   // the same network as SCL:
   "Carrier_58_Carrier_In_Zone" := "EMS".Carrier[58].SDC_OUT.Zone;
END_REGION
